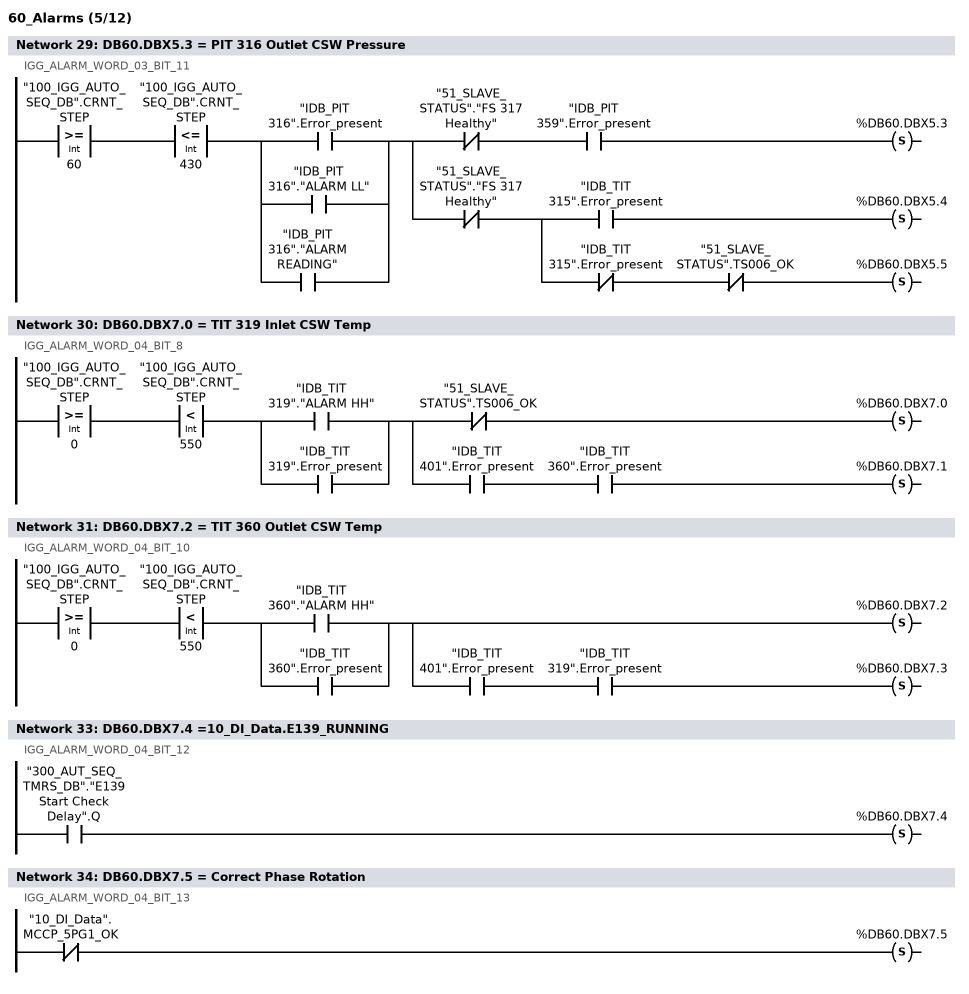
   RUNG wire#powerrail
      { S7_Templates := "SrcType := Int" } GE_Contact(in1 := "100_IGG_AUTO_SEQ_DB".CRNT_STEP, in2 := 60)
      { S7_Templates := "SrcType := Int" } LE_Contact(in1 := "100_IGG_AUTO_SEQ_DB".CRNT_STEP, in2 := 430)
      wire#w1
      Contact( "IDB_PIT 316".Error_present )
      wire#w2
      I_Contact( "51_SLAVE_STATUS"."FS 317 Healthy" )
      Contact( "IDB_PIT 359".Error_present )
      S_Coil( %DB60.DBX5.3 )
   END_RUNG
   RUNG wire#w1
      Contact( "IDB_PIT 316"."ALARM LL" )
   END_RUNG wire#w2
   RUNG wire#w1
      Contact( "IDB_PIT 316"."ALARM READING" )
   END_RUNG wire#w2
   RUNG wire#w2
      I_Contact( "51_SLAVE_STATUS"."FS 317 Healthy" )
      wire#w3
      Contact( "IDB_TIT 315".Error_present )
      S_Coil( %DB60.DBX5.4 )
   END_RUNG
   RUNG wire#w3
      I_Contact( "IDB_TIT 315".Error_present )
      I_Contact( "51_SLAVE_STATUS".TS006_OK )
      S_Coil( %DB60.DBX5.5 )
   END_RUNG
   // the same network as SCL:
   #_w1 := ("100_IGG_AUTO_SEQ_DB".CRNT_STEP >= 60) AND ("100_IGG_AUTO_SEQ_DB".CRNT_STEP <= 430) AND ("IDB_PIT 316".Error_present OR "IDB_PIT 316"."ALARM LL" OR "IDB_PIT 316"."ALARM READING");
   IF #_w1 AND NOT "51_SLAVE_STATUS"."FS 317 Healthy" AND "IDB_PIT 359".Error_present THEN
       %DB60.DBX5.3 := TRUE;
   END_IF;
   #_w2 := #_w1 AND NOT "51_SLAVE_STATUS"."FS 317 Healthy";
   IF #_w2 AND "IDB_TIT 315".Error_present THEN %DB60.DBX5.4 := TRUE; END_IF;
   IF #_w2 AND NOT "IDB_TIT 315".Error_present AND NOT "51_SLAVE_STATUS".TS006_OK THEN
       %DB60.DBX5.5 := TRUE;
   END_IF;
END_REGION

REGION Network 30: DB60.DBX7.0 = TIT 319 Inlet CSW Temp
   // IGG_ALARM_WORD_04_BIT_8
   RUNG wire#powerrail
      { S7_Templates := "SrcType := Int" } GE_Contact(in1 := "100_IGG_AUTO_SEQ_DB".CRNT_STEP, in2 := 0)
      { S7_Templates := "SrcType := Int" } LT_Contact(in1 := "100_IGG_AUTO_SEQ_DB".CRNT_STEP, in2 := 550)
      wire#w1
      Contact( "IDB_TIT 319"."ALARM HH" )
      wire#w2
      I_Contact( "51_SLAVE_STATUS".TS006_OK )
      S_Coil( %DB60.DBX7.0 )
   END_RUNG
   RUNG wire#w1
      Contact( "IDB_TIT 319".Error_present )
   END_RUNG wire#w2
   RUNG wire#w2
      Contact( "IDB_TIT 401".Error_present )
      Contact( "IDB_TIT 360".Error_present )
      S_Coil( %DB60.DBX7.1 )
   END_RUNG
   // the same network as SCL:
   #_w1 := ("100_IGG_AUTO_SEQ_DB".CRNT_STEP >= 0) AND ("100_IGG_AUTO_SEQ_DB".CRNT_STEP < 550) AND ("IDB_TIT 319"."ALARM HH" OR "IDB_TIT 319".Error_present);
   IF #_w1 AND NOT "51_SLAVE_STATUS".TS006_OK THEN %DB60.DBX7.0 := TRUE; END_IF;
   IF #_w1 AND "IDB_TIT 401".Error_present AND "IDB_TIT 360".Error_present THEN %DB60.DBX7.1 := TRUE; END_IF;
END_REGION

REGION Network 31: DB60.DBX7.2 = TIT 360 Outlet CSW Temp
   // IGG_ALARM_WORD_04_BIT_10
   RUNG wire#powerrail
      { S7_Templates := "SrcType := Int" } GE_Contact(in1 := "100_IGG_AUTO_SEQ_DB".CRNT_STEP, in2 := 0)
      { S7_Templates := "SrcType := Int" } LT_Contact(in1 := "100_IGG_AUTO_SEQ_DB".CRNT_STEP, in2 := 550)
      wire#w1
      Contact( "IDB_TIT 360"."ALARM HH" )
      wire#w2
      S_Coil( %DB60.DBX7.2 )
   END_RUNG
   RUNG wire#w1
      Contact( "IDB_TIT 360".Error_present )
   END_RUNG wire#w2
   RUNG wire#w2
      Contact( "IDB_TIT 401".Error_present )
      Contact( "IDB_TIT 319".Error_present )
      S_Coil( %DB60.DBX7.3 )
   END_RUNG
   // the same network as SCL:
   #_w1 := ("100_IGG_AUTO_SEQ_DB".CRNT_STEP >= 0) AND ("100_IGG_AUTO_SEQ_DB".CRNT_STEP < 550) AND ("IDB_TIT 360"."ALARM HH" OR "IDB_TIT 360".Error_present);
   IF #_w1 THEN %DB60.DBX7.2 := TRUE; END_IF;
   IF #_w1 AND "IDB_TIT 401".Error_present AND "IDB_TIT 319".Error_present THEN %DB60.DBX7.3 := TRUE; END_IF;
END_REGION

REGION Network 33: DB60.DBX7.4 =10_DI_Data.E139_RUNNING
   // IGG_ALARM_WORD_04_BIT_12
   RUNG wire#powerrail
      Contact( "300_AUT_SEQ_TMRS_DB"."E139 Start Check Delay".Q )
      S_Coil( %DB60.DBX7.4 )
   END_RUNG
   // the same network as SCL:
   IF "300_AUT_SEQ_TMRS_DB"."E139 Start Check Delay".Q THEN %DB60.DBX7.4 := TRUE; END_IF;
END_REGION

REGION Network 34: DB60.DBX7.5 = Correct Phase Rotation
   // IGG_ALARM_WORD_04_BIT_13
   RUNG wire#powerrail
      I_Contact( "10_DI_Data".MCCP_5PG1_OK )
      S_Coil( %DB60.DBX7.5 )
   END_RUNG
   // the same network as SCL:
   IF NOT "10_DI_Data".MCCP_5PG1_OK THEN %DB60.DBX7.5 := TRUE; END_IF;
END_REGION

REGION Network 36: DB60.DBX6.0 = CV311 Fault
   // IGG_ALARM_WORD_04_BIT_0
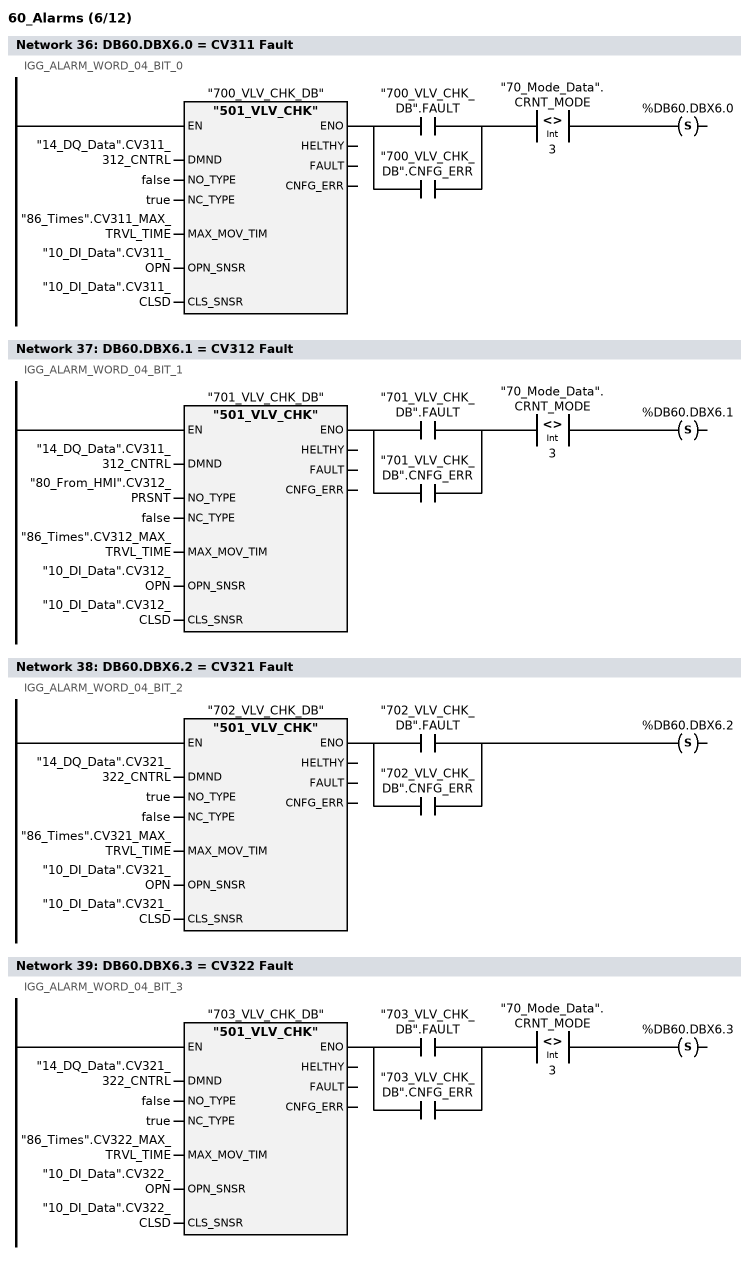
   RUNG wire#powerrail
      "700_VLV_CHK_DB"(DMND := "14_DQ_Data".CV311_312_CNTRL, NO_TYPE := false, NC_TYPE := true, MAX_MOV_TIM := "86_Times".CV311_MAX_TRVL_TIME, OPN_SNSR := "10_DI_Data".CV311_OPN, CLS_SNSR := "10_DI_Data".CV311_CLSD, HELTHY =>, FAULT =>, CNFG_ERR =>)
      wire#w1
      Contact( "700_VLV_CHK_DB".FAULT )
      wire#w2
      { S7_Templates := "SrcType := Int" } NE_Contact(in1 := "70_Mode_Data".CRNT_MODE, in2 := 3)
      S_Coil( %DB60.DBX6.0 )
   END_RUNG
   RUNG wire#w1
      Contact( "700_VLV_CHK_DB".CNFG_ERR )
   END_RUNG wire#w2
   // the same network as SCL:
   "700_VLV_CHK_DB"(DMND := "14_DQ_Data".CV311_312_CNTRL,   // "501_VLV_CHK"
                    NO_TYPE := false,
                    NC_TYPE := true,
                    MAX_MOV_TIM := "86_Times".CV311_MAX_TRVL_TIME,
                    OPN_SNSR := "10_DI_Data".CV311_OPN,
                    CLS_SNSR := "10_DI_Data".CV311_CLSD,
                    ENO => #_w1);
   IF #_w1 AND ("700_VLV_CHK_DB".FAULT OR "700_VLV_CHK_DB".CNFG_ERR) AND ("70_Mode_Data".CRNT_MODE <> 3) THEN
       %DB60.DBX6.0 := TRUE;
   END_IF;
END_REGION

REGION Network 37: DB60.DBX6.1 = CV312 Fault
   // IGG_ALARM_WORD_04_BIT_1
   RUNG wire#powerrail
      "701_VLV_CHK_DB"(DMND := "14_DQ_Data".CV311_312_CNTRL, NO_TYPE := "80_From_HMI".CV312_PRSNT, NC_TYPE := false, MAX_MOV_TIM := "86_Times".CV312_MAX_TRVL_TIME, OPN_SNSR := "10_DI_Data".CV312_OPN, CLS_SNSR := "10_DI_Data".CV312_CLSD, HELTHY =>, FAULT =>, CNFG_ERR =>)
      wire#w1
      Contact( "701_VLV_CHK_DB".FAULT )
      wire#w2
      { S7_Templates := "SrcType := Int" } NE_Contact(in1 := "70_Mode_Data".CRNT_MODE, in2 := 3)
      S_Coil( %DB60.DBX6.1 )
   END_RUNG
   RUNG wire#w1
      Contact( "701_VLV_CHK_DB".CNFG_ERR )
   END_RUNG wire#w2
   // the same network as SCL:
   "701_VLV_CHK_DB"(DMND := "14_DQ_Data".CV311_312_CNTRL,   // "501_VLV_CHK"
                    NO_TYPE := "80_From_HMI".CV312_PRSNT,
                    NC_TYPE := false,
                    MAX_MOV_TIM := "86_Times".CV312_MAX_TRVL_TIME,
                    OPN_SNSR := "10_DI_Data".CV312_OPN,
                    CLS_SNSR := "10_DI_Data".CV312_CLSD,
                    ENO => #_w1);
   IF #_w1 AND ("701_VLV_CHK_DB".FAULT OR "701_VLV_CHK_DB".CNFG_ERR) AND ("70_Mode_Data".CRNT_MODE <> 3) THEN
       %DB60.DBX6.1 := TRUE;
   END_IF;
END_REGION

REGION Network 38: DB60.DBX6.2 = CV321 Fault
   // IGG_ALARM_WORD_04_BIT_2
   RUNG wire#powerrail
      "702_VLV_CHK_DB"(DMND := "14_DQ_Data".CV321_322_CNTRL, NO_TYPE := true, NC_TYPE := false, MAX_MOV_TIM := "86_Times".CV321_MAX_TRVL_TIME, OPN_SNSR := "10_DI_Data".CV321_OPN, CLS_SNSR := "10_DI_Data".CV321_CLSD, HELTHY =>, FAULT =>, CNFG_ERR =>)
      wire#w1
      Contact( "702_VLV_CHK_DB".FAULT )
      wire#w2
      S_Coil( %DB60.DBX6.2 )
   END_RUNG
   RUNG wire#w1
      Contact( "702_VLV_CHK_DB".CNFG_ERR )
   END_RUNG wire#w2
   // the same network as SCL:
   "702_VLV_CHK_DB"(DMND := "14_DQ_Data".CV321_322_CNTRL,   // "501_VLV_CHK"
                    NO_TYPE := true,
                    NC_TYPE := false,
                    MAX_MOV_TIM := "86_Times".CV321_MAX_TRVL_TIME,
                    OPN_SNSR := "10_DI_Data".CV321_OPN,
                    CLS_SNSR := "10_DI_Data".CV321_CLSD,
                    ENO => #_w1);
   IF #_w1 AND ("702_VLV_CHK_DB".FAULT OR "702_VLV_CHK_DB".CNFG_ERR) THEN %DB60.DBX6.2 := TRUE; END_IF;
END_REGION

REGION Network 39: DB60.DBX6.3 = CV322 Fault
   // IGG_ALARM_WORD_04_BIT_3
   RUNG wire#powerrail
      "703_VLV_CHK_DB"(DMND := "14_DQ_Data".CV321_322_CNTRL, NO_TYPE := false, NC_TYPE := true, MAX_MOV_TIM := "86_Times".CV322_MAX_TRVL_TIME, OPN_SNSR := "10_DI_Data".CV322_OPN, CLS_SNSR := "10_DI_Data".CV322_CLSD, HELTHY =>, FAULT =>, CNFG_ERR =>)
      wire#w1
      Contact( "703_VLV_CHK_DB".FAULT )
      wire#w2
      { S7_Templates := "SrcType := Int" } NE_Contact(in1 := "70_Mode_Data".CRNT_MODE, in2 := 3)
      S_Coil( %DB60.DBX6.3 )
   END_RUNG
   RUNG wire#w1
      Contact( "703_VLV_CHK_DB".CNFG_ERR )
   END_RUNG wire#w2
   // the same network as SCL:
   "703_VLV_CHK_DB"(DMND := "14_DQ_Data".CV321_322_CNTRL,   // "501_VLV_CHK"
                    NO_TYPE := false,
                    NC_TYPE := true,
                    MAX_MOV_TIM := "86_Times".CV322_MAX_TRVL_TIME,
                    OPN_SNSR := "10_DI_Data".CV322_OPN,
                    CLS_SNSR := "10_DI_Data".CV322_CLSD,
                    ENO => #_w1);
   IF #_w1 AND ("703_VLV_CHK_DB".FAULT OR "703_VLV_CHK_DB".CNFG_ERR) AND ("70_Mode_Data".CRNT_MODE <> 3) THEN
       %DB60.DBX6.3 := TRUE;
   END_IF;
END_REGION

REGION Network 40: DB60.DBX6.4 = CV401 Fault
   // IGG_ALARM_WORD_04_BIT_4
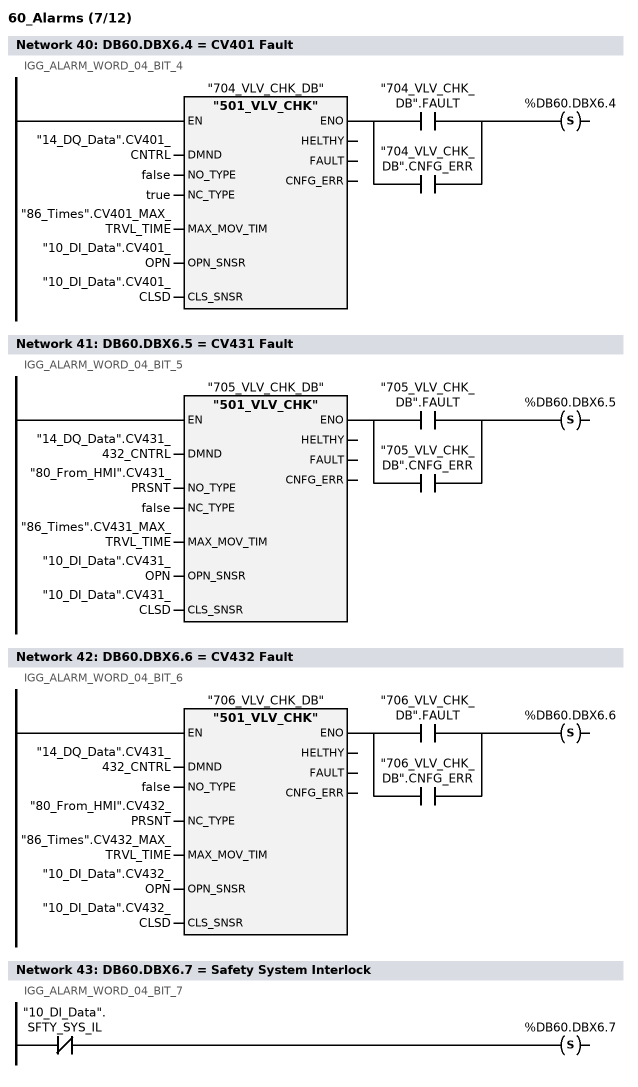
   RUNG wire#powerrail
      "704_VLV_CHK_DB"(DMND := "14_DQ_Data".CV401_CNTRL, NO_TYPE := false, NC_TYPE := true, MAX_MOV_TIM := "86_Times".CV401_MAX_TRVL_TIME, OPN_SNSR := "10_DI_Data".CV401_OPN, CLS_SNSR := "10_DI_Data".CV401_CLSD, HELTHY =>, FAULT =>, CNFG_ERR =>)
      wire#w1
      Contact( "704_VLV_CHK_DB".FAULT )
      wire#w2
      S_Coil( %DB60.DBX6.4 )
   END_RUNG
   RUNG wire#w1
      Contact( "704_VLV_CHK_DB".CNFG_ERR )
   END_RUNG wire#w2
   // the same network as SCL:
   "704_VLV_CHK_DB"(DMND := "14_DQ_Data".CV401_CNTRL,   // "501_VLV_CHK"
                    NO_TYPE := false,
                    NC_TYPE := true,
                    MAX_MOV_TIM := "86_Times".CV401_MAX_TRVL_TIME,
                    OPN_SNSR := "10_DI_Data".CV401_OPN,
                    CLS_SNSR := "10_DI_Data".CV401_CLSD,
                    ENO => #_w1);
   IF #_w1 AND ("704_VLV_CHK_DB".FAULT OR "704_VLV_CHK_DB".CNFG_ERR) THEN %DB60.DBX6.4 := TRUE; END_IF;
END_REGION

REGION Network 41: DB60.DBX6.5 = CV431 Fault
   // IGG_ALARM_WORD_04_BIT_5
   RUNG wire#powerrail
      "705_VLV_CHK_DB"(DMND := "14_DQ_Data".CV431_432_CNTRL, NO_TYPE := "80_From_HMI".CV431_PRSNT, NC_TYPE := false, MAX_MOV_TIM := "86_Times".CV431_MAX_TRVL_TIME, OPN_SNSR := "10_DI_Data".CV431_OPN, CLS_SNSR := "10_DI_Data".CV431_CLSD, HELTHY =>, FAULT =>, CNFG_ERR =>)
      wire#w1
      Contact( "705_VLV_CHK_DB".FAULT )
      wire#w2
      S_Coil( %DB60.DBX6.5 )
   END_RUNG
   RUNG wire#w1
      Contact( "705_VLV_CHK_DB".CNFG_ERR )
   END_RUNG wire#w2
   // the same network as SCL:
   "705_VLV_CHK_DB"(DMND := "14_DQ_Data".CV431_432_CNTRL,   // "501_VLV_CHK"
                    NO_TYPE := "80_From_HMI".CV431_PRSNT,
                    NC_TYPE := false,
                    MAX_MOV_TIM := "86_Times".CV431_MAX_TRVL_TIME,
                    OPN_SNSR := "10_DI_Data".CV431_OPN,
                    CLS_SNSR := "10_DI_Data".CV431_CLSD,
                    ENO => #_w1);
   IF #_w1 AND ("705_VLV_CHK_DB".FAULT OR "705_VLV_CHK_DB".CNFG_ERR) THEN %DB60.DBX6.5 := TRUE; END_IF;
END_REGION

REGION Network 42: DB60.DBX6.6 = CV432 Fault
   // IGG_ALARM_WORD_04_BIT_6
   RUNG wire#powerrail
      "706_VLV_CHK_DB"(DMND := "14_DQ_Data".CV431_432_CNTRL, NO_TYPE := false, NC_TYPE := "80_From_HMI".CV432_PRSNT, MAX_MOV_TIM := "86_Times".CV432_MAX_TRVL_TIME, OPN_SNSR := "10_DI_Data".CV432_OPN, CLS_SNSR := "10_DI_Data".CV432_CLSD, HELTHY =>, FAULT =>, CNFG_ERR =>)
      wire#w1
      Contact( "706_VLV_CHK_DB".FAULT )
      wire#w2
      S_Coil( %DB60.DBX6.6 )
   END_RUNG
   RUNG wire#w1
      Contact( "706_VLV_CHK_DB".CNFG_ERR )
   END_RUNG wire#w2
   // the same network as SCL:
   "706_VLV_CHK_DB"(DMND := "14_DQ_Data".CV431_432_CNTRL,   // "501_VLV_CHK"
                    NO_TYPE := false,
                    NC_TYPE := "80_From_HMI".CV432_PRSNT,
                    MAX_MOV_TIM := "86_Times".CV432_MAX_TRVL_TIME,
                    OPN_SNSR := "10_DI_Data".CV432_OPN,
                    CLS_SNSR := "10_DI_Data".CV432_CLSD,
                    ENO => #_w1);
   IF #_w1 AND ("706_VLV_CHK_DB".FAULT OR "706_VLV_CHK_DB".CNFG_ERR) THEN %DB60.DBX6.6 := TRUE; END_IF;
END_REGION

REGION Network 43: DB60.DBX6.7 = Safety System Interlock
   // IGG_ALARM_WORD_04_BIT_7
   RUNG wire#powerrail
      I_Contact( "10_DI_Data".SFTY_SYS_IL )
      S_Coil( %DB60.DBX6.7 )
   END_RUNG
   // the same network as SCL:
   IF NOT "10_DI_Data".SFTY_SYS_IL THEN %DB60.DBX6.7 := TRUE; END_IF;
END_REGION

REGION Network 45: New Alarm Check
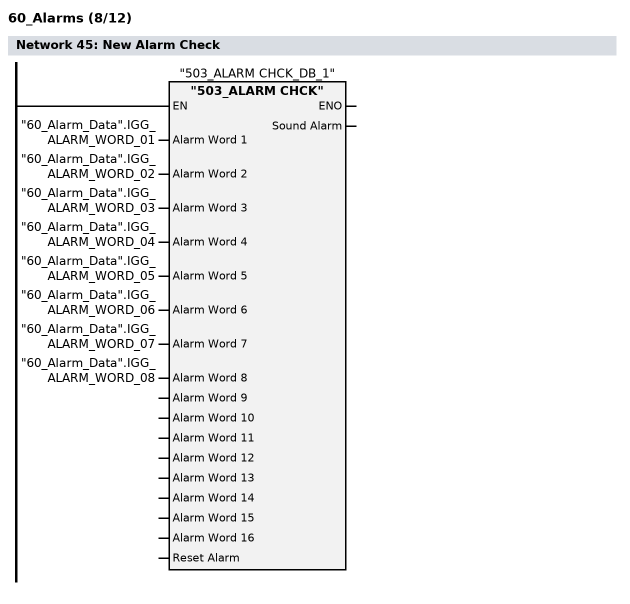
   RUNG wire#powerrail
      "503_ALARM CHCK_DB_1"("Alarm Word 1" := "60_Alarm_Data".IGG_ALARM_WORD_01, "Alarm Word 2" := "60_Alarm_Data".IGG_ALARM_WORD_02, "Alarm Word 3" := "60_Alarm_Data".IGG_ALARM_WORD_03, "Alarm Word 4" := "60_Alarm_Data".IGG_ALARM_WORD_04, "Alarm Word 5" := "60_Alarm_Data".IGG_ALARM_WORD_05, "Alarm Word 6" := "60_Alarm_Data".IGG_ALARM_WORD_06, "Alarm Word 7" := "60_Alarm_Data".IGG_ALARM_WORD_07, "Alarm Word 8" := "60_Alarm_Data".IGG_ALARM_WORD_08, "Alarm Word 9" :=, "Alarm Word 10" :=, "Alarm Word 11" :=, "Alarm Word 12" :=, "Alarm Word 13" :=, "Alarm Word 14" :=, "Alarm Word 15" :=, "Alarm Word 16" :=, "Reset Alarm" :=, "Sound Alarm" =>)
   END_RUNG
   // the same network as SCL:
   "503_ALARM CHCK_DB_1"("Alarm Word 1" := "60_Alarm_Data".IGG_ALARM_WORD_01,   // "503_ALARM CHCK"
                         "Alarm Word 2" := "60_Alarm_Data".IGG_ALARM_WORD_02,
                         "Alarm Word 3" := "60_Alarm_Data".IGG_ALARM_WORD_03,
                         "Alarm Word 4" := "60_Alarm_Data".IGG_ALARM_WORD_04,
                         "Alarm Word 5" := "60_Alarm_Data".IGG_ALARM_WORD_05,
                         "Alarm Word 6" := "60_Alarm_Data".IGG_ALARM_WORD_06,
                         "Alarm Word 7" := "60_Alarm_Data".IGG_ALARM_WORD_07,
                         "Alarm Word 8" := "60_Alarm_Data".IGG_ALARM_WORD_08);
END_REGION

REGION Network 46: Alarm reset
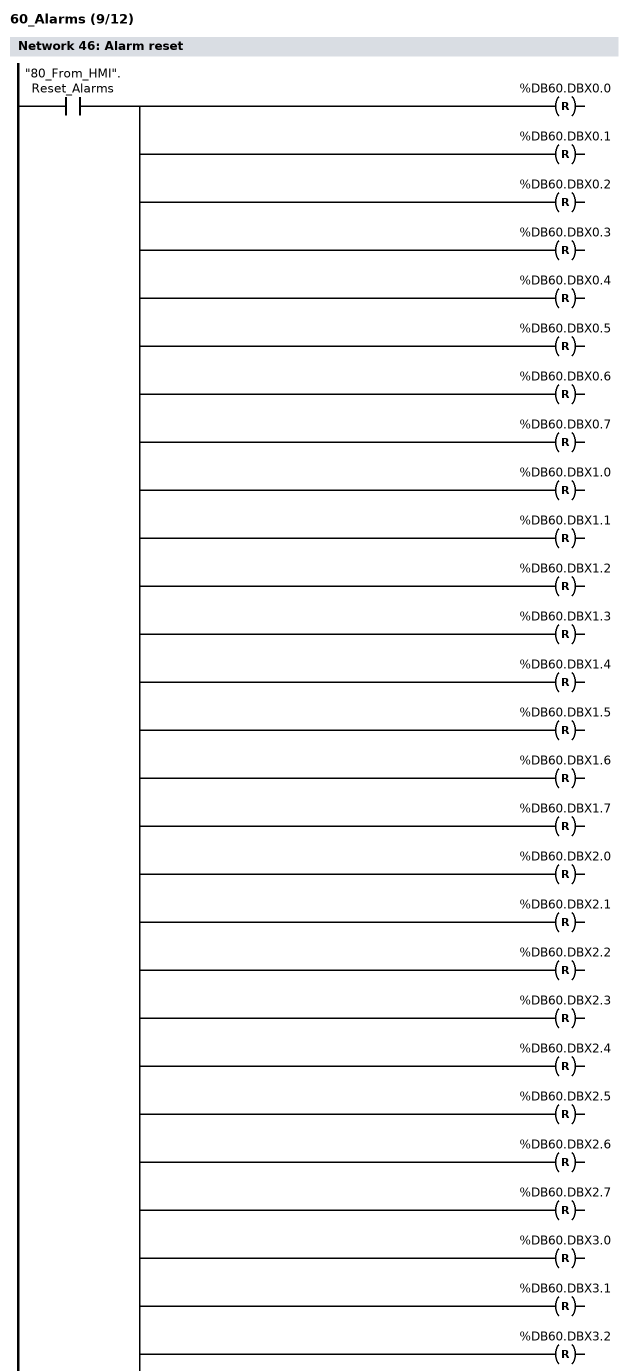
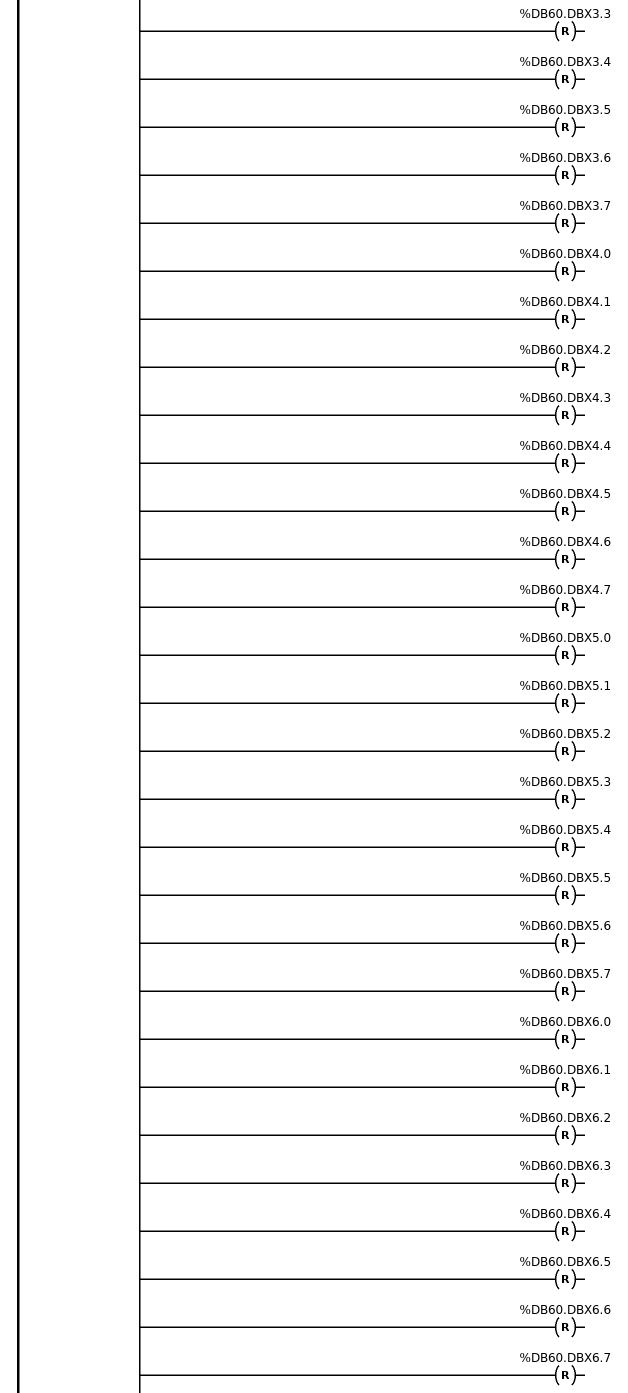
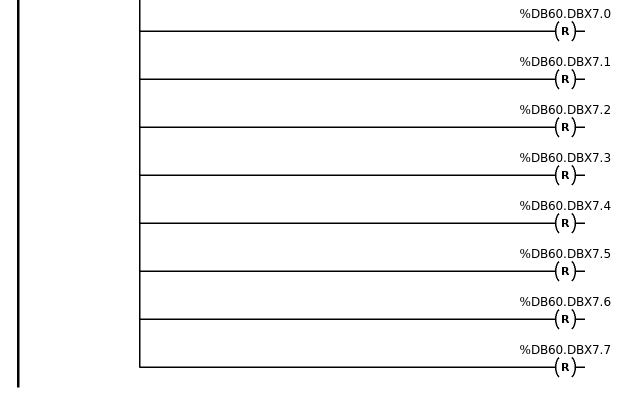
   RUNG wire#powerrail
      Contact( "80_From_HMI".Reset_Alarms )
      wire#w1
      R_Coil( %DB60.DBX0.0 )
   END_RUNG
   RUNG wire#w1
      R_Coil( %DB60.DBX0.1 )
   END_RUNG
   RUNG wire#w1
      R_Coil( %DB60.DBX0.2 )
   END_RUNG
   RUNG wire#w1
      R_Coil( %DB60.DBX0.3 )
   END_RUNG
   RUNG wire#w1
      R_Coil( %DB60.DBX0.4 )
   END_RUNG
   RUNG wire#w1
      R_Coil( %DB60.DBX0.5 )
   END_RUNG
   RUNG wire#w1
      R_Coil( %DB60.DBX0.6 )
   END_RUNG
   RUNG wire#w1
      R_Coil( %DB60.DBX0.7 )
   END_RUNG
   RUNG wire#w1
      R_Coil( %DB60.DBX1.0 )
   END_RUNG
   RUNG wire#w1
      R_Coil( %DB60.DBX1.1 )
   END_RUNG
   RUNG wire#w1
      R_Coil( %DB60.DBX1.2 )
   END_RUNG
   RUNG wire#w1
      R_Coil( %DB60.DBX1.3 )
   END_RUNG
   RUNG wire#w1
      R_Coil( %DB60.DBX1.4 )
   END_RUNG
   RUNG wire#w1
      R_Coil( %DB60.DBX1.5 )
   END_RUNG
   RUNG wire#w1
      R_Coil( %DB60.DBX1.6 )
   END_RUNG
   RUNG wire#w1
      R_Coil( %DB60.DBX1.7 )
   END_RUNG
   RUNG wire#w1
      R_Coil( %DB60.DBX2.0 )
   END_RUNG
   RUNG wire#w1
      R_Coil( %DB60.DBX2.1 )
   END_RUNG
   RUNG wire#w1
      R_Coil( %DB60.DBX2.2 )
   END_RUNG
   RUNG wire#w1
      R_Coil( %DB60.DBX2.3 )
   END_RUNG
   RUNG wire#w1
      R_Coil( %DB60.DBX2.4 )
   END_RUNG
   RUNG wire#w1
      R_Coil( %DB60.DBX2.5 )
   END_RUNG
   RUNG wire#w1
      R_Coil( %DB60.DBX2.6 )
   END_RUNG
   RUNG wire#w1
      R_Coil( %DB60.DBX2.7 )
   END_RUNG
   RUNG wire#w1
      R_Coil( %DB60.DBX3.0 )
   END_RUNG
   RUNG wire#w1
      R_Coil( %DB60.DBX3.1 )
   END_RUNG
   RUNG wire#w1
      R_Coil( %DB60.DBX3.2 )
   END_RUNG
   RUNG wire#w1
      R_Coil( %DB60.DBX3.3 )
   END_RUNG
   RUNG wire#w1
      R_Coil( %DB60.DBX3.4 )
   END_RUNG
   RUNG wire#w1
      R_Coil( %DB60.DBX3.5 )
   END_RUNG
   RUNG wire#w1
      R_Coil( %DB60.DBX3.6 )
   END_RUNG
   RUNG wire#w1
      R_Coil( %DB60.DBX3.7 )
   END_RUNG
   RUNG wire#w1
      R_Coil( %DB60.DBX4.0 )
   END_RUNG
   RUNG wire#w1
      R_Coil( %DB60.DBX4.1 )
   END_RUNG
   RUNG wire#w1
      R_Coil( %DB60.DBX4.2 )
   END_RUNG
   RUNG wire#w1
      R_Coil( %DB60.DBX4.3 )
   END_RUNG
   RUNG wire#w1
      R_Coil( %DB60.DBX4.4 )
   END_RUNG
   RUNG wire#w1
      R_Coil( %DB60.DBX4.5 )
   END_RUNG
   RUNG wire#w1
      R_Coil( %DB60.DBX4.6 )
   END_RUNG
   RUNG wire#w1
      R_Coil( %DB60.DBX4.7 )
   END_RUNG
   RUNG wire#w1
      R_Coil( %DB60.DBX5.0 )
   END_RUNG
   RUNG wire#w1
      R_Coil( %DB60.DBX5.1 )
   END_RUNG
   RUNG wire#w1
      R_Coil( %DB60.DBX5.2 )
   END_RUNG
   RUNG wire#w1
      R_Coil( %DB60.DBX5.3 )
   END_RUNG
   RUNG wire#w1
      R_Coil( %DB60.DBX5.4 )
   END_RUNG
   RUNG wire#w1
      R_Coil( %DB60.DBX5.5 )
   END_RUNG
   RUNG wire#w1
      R_Coil( %DB60.DBX5.6 )
   END_RUNG
   RUNG wire#w1
      R_Coil( %DB60.DBX5.7 )
   END_RUNG
   RUNG wire#w1
      R_Coil( %DB60.DBX6.0 )
   END_RUNG
   RUNG wire#w1
      R_Coil( %DB60.DBX6.1 )
   END_RUNG
   RUNG wire#w1
      R_Coil( %DB60.DBX6.2 )
   END_RUNG
   RUNG wire#w1
      R_Coil( %DB60.DBX6.3 )
   END_RUNG
   RUNG wire#w1
      R_Coil( %DB60.DBX6.4 )
   END_RUNG
   RUNG wire#w1
      R_Coil( %DB60.DBX6.5 )
   END_RUNG
   RUNG wire#w1
      R_Coil( %DB60.DBX6.6 )
   END_RUNG
   RUNG wire#w1
      R_Coil( %DB60.DBX6.7 )
   END_RUNG
   RUNG wire#w1
      R_Coil( %DB60.DBX7.0 )
   END_RUNG
   RUNG wire#w1
      R_Coil( %DB60.DBX7.1 )
   END_RUNG
   RUNG wire#w1
      R_Coil( %DB60.DBX7.2 )
   END_RUNG
   RUNG wire#w1
      R_Coil( %DB60.DBX7.3 )
   END_RUNG
   RUNG wire#w1
      R_Coil( %DB60.DBX7.4 )
   END_RUNG
   RUNG wire#w1
      R_Coil( %DB60.DBX7.5 )
   END_RUNG
   RUNG wire#w1
      R_Coil( %DB60.DBX7.6 )
   END_RUNG
   RUNG wire#w1
      R_Coil( %DB60.DBX7.7 )
   END_RUNG
   // the same network as SCL:
   IF "80_From_HMI".Reset_Alarms THEN
       %DB60.DBX0.0 := FALSE;
       %DB60.DBX0.1 := FALSE;
       %DB60.DBX0.2 := FALSE;
       %DB60.DBX0.3 := FALSE;
       %DB60.DBX0.4 := FALSE;
       %DB60.DBX0.5 := FALSE;
       %DB60.DBX0.6 := FALSE;
       %DB60.DBX0.7 := FALSE;
       %DB60.DBX1.0 := FALSE;
       %DB60.DBX1.1 := FALSE;
       %DB60.DBX1.2 := FALSE;
       %DB60.DBX1.3 := FALSE;
       %DB60.DBX1.4 := FALSE;
       %DB60.DBX1.5 := FALSE;
       %DB60.DBX1.6 := FALSE;
       %DB60.DBX1.7 := FALSE;
       %DB60.DBX2.0 := FALSE;
       %DB60.DBX2.1 := FALSE;
       %DB60.DBX2.2 := FALSE;
       %DB60.DBX2.3 := FALSE;
       %DB60.DBX2.4 := FALSE;
       %DB60.DBX2.5 := FALSE;
       %DB60.DBX2.6 := FALSE;
       %DB60.DBX2.7 := FALSE;
       %DB60.DBX3.0 := FALSE;
       %DB60.DBX3.1 := FALSE;
       %DB60.DBX3.2 := FALSE;
       %DB60.DBX3.3 := FALSE;
       %DB60.DBX3.4 := FALSE;
       %DB60.DBX3.5 := FALSE;
       %DB60.DBX3.6 := FALSE;
       %DB60.DBX3.7 := FALSE;
       %DB60.DBX4.0 := FALSE;
       %DB60.DBX4.1 := FALSE;
       %DB60.DBX4.2 := FALSE;
       %DB60.DBX4.3 := FALSE;
       %DB60.DBX4.4 := FALSE;
       %DB60.DBX4.5 := FALSE;
       %DB60.DBX4.6 := FALSE;
       %DB60.DBX4.7 := FALSE;
       %DB60.DBX5.0 := FALSE;
       %DB60.DBX5.1 := FALSE;
       %DB60.DBX5.2 := FALSE;
       %DB60.DBX5.3 := FALSE;
       %DB60.DBX5.4 := FALSE;
       %DB60.DBX5.5 := FALSE;
       %DB60.DBX5.6 := FALSE;
       %DB60.DBX5.7 := FALSE;
       %DB60.DBX6.0 := FALSE;
       %DB60.DBX6.1 := FALSE;
       %DB60.DBX6.2 := FALSE;
       %DB60.DBX6.3 := FALSE;
       %DB60.DBX6.4 := FALSE;
       %DB60.DBX6.5 := FALSE;
       %DB60.DBX6.6 := FALSE;
       %DB60.DBX6.7 := FALSE;
       %DB60.DBX7.0 := FALSE;
       %DB60.DBX7.1 := FALSE;
       %DB60.DBX7.2 := FALSE;
       %DB60.DBX7.3 := FALSE;
       %DB60.DBX7.4 := FALSE;
       %DB60.DBX7.5 := FALSE;
       %DB60.DBX7.6 := FALSE;
       %DB60.DBX7.7 := FALSE;
   END_IF;
END_REGION

REGION Network 47: Alarm reset II
   // testing
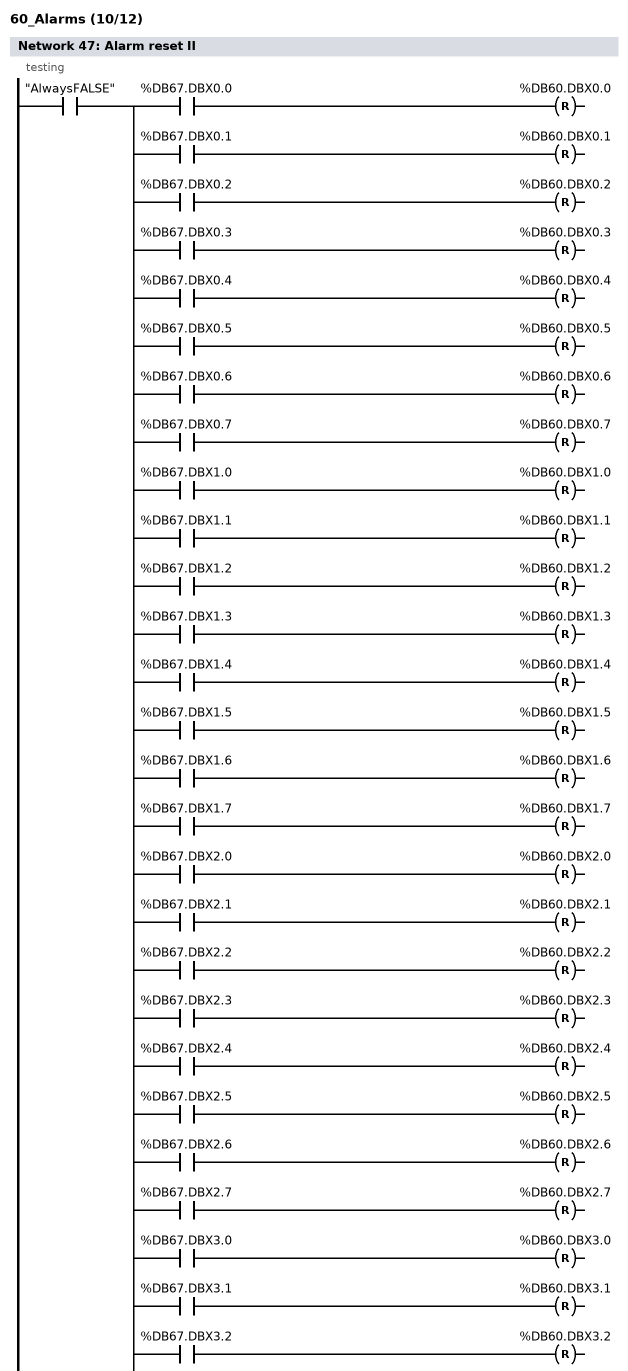
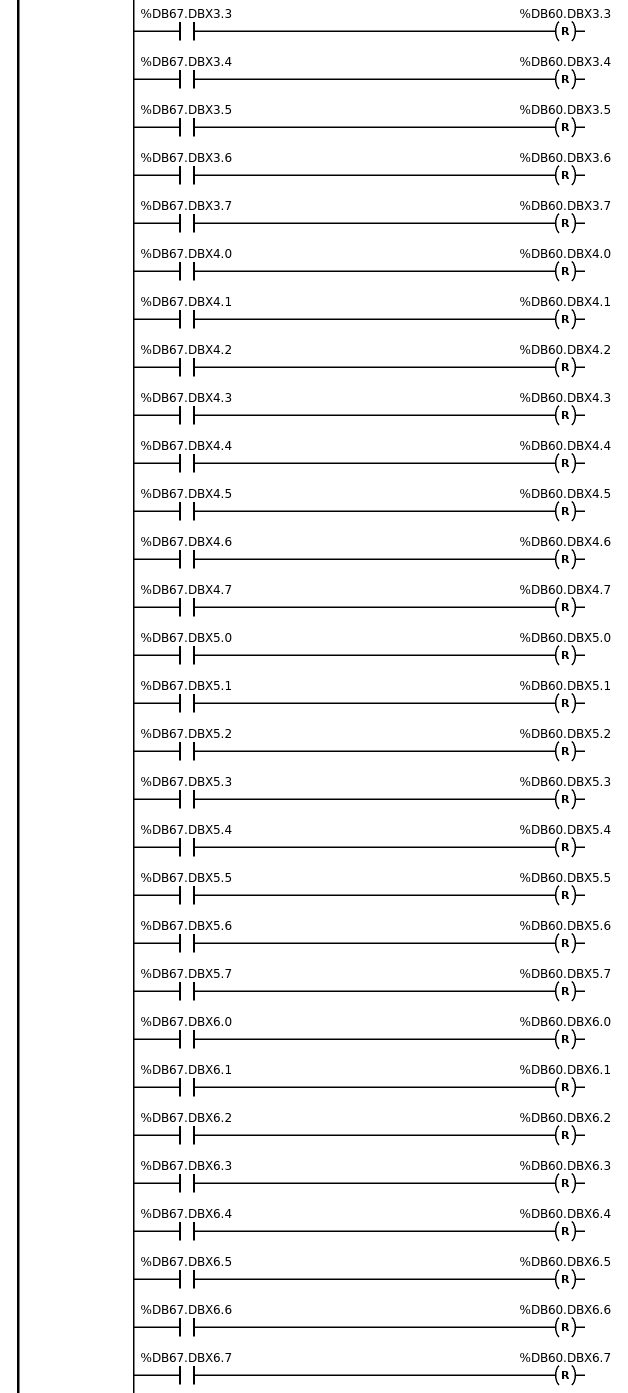
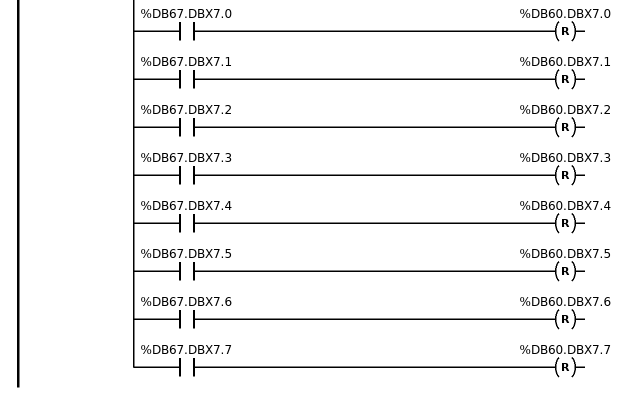
   RUNG wire#powerrail
      Contact( "AlwaysFALSE" )
      wire#w1
      Contact( %DB67.DBX0.0 )
      R_Coil( %DB60.DBX0.0 )
   END_RUNG
   RUNG wire#w1
      Contact( %DB67.DBX0.1 )
      R_Coil( %DB60.DBX0.1 )
   END_RUNG
   RUNG wire#w1
      Contact( %DB67.DBX0.2 )
      R_Coil( %DB60.DBX0.2 )
   END_RUNG
   RUNG wire#w1
      Contact( %DB67.DBX0.3 )
      R_Coil( %DB60.DBX0.3 )
   END_RUNG
   RUNG wire#w1
      Contact( %DB67.DBX0.4 )
      R_Coil( %DB60.DBX0.4 )
   END_RUNG
   RUNG wire#w1
      Contact( %DB67.DBX0.5 )
      R_Coil( %DB60.DBX0.5 )
   END_RUNG
   RUNG wire#w1
      Contact( %DB67.DBX0.6 )
      R_Coil( %DB60.DBX0.6 )
   END_RUNG
   RUNG wire#w1
      Contact( %DB67.DBX0.7 )
      R_Coil( %DB60.DBX0.7 )
   END_RUNG
   RUNG wire#w1
      Contact( %DB67.DBX1.0 )
      R_Coil( %DB60.DBX1.0 )
   END_RUNG
   RUNG wire#w1
      Contact( %DB67.DBX1.1 )
      R_Coil( %DB60.DBX1.1 )
   END_RUNG
   RUNG wire#w1
      Contact( %DB67.DBX1.2 )
      R_Coil( %DB60.DBX1.2 )
   END_RUNG
   RUNG wire#w1
      Contact( %DB67.DBX1.3 )
      R_Coil( %DB60.DBX1.3 )
   END_RUNG
   RUNG wire#w1
      Contact( %DB67.DBX1.4 )
      R_Coil( %DB60.DBX1.4 )
   END_RUNG
   RUNG wire#w1
      Contact( %DB67.DBX1.5 )
      R_Coil( %DB60.DBX1.5 )
   END_RUNG
   RUNG wire#w1
      Contact( %DB67.DBX1.6 )
      R_Coil( %DB60.DBX1.6 )
   END_RUNG
   RUNG wire#w1
      Contact( %DB67.DBX1.7 )
      R_Coil( %DB60.DBX1.7 )
   END_RUNG
   RUNG wire#w1
      Contact( %DB67.DBX2.0 )
      R_Coil( %DB60.DBX2.0 )
   END_RUNG
   RUNG wire#w1
      Contact( %DB67.DBX2.1 )
      R_Coil( %DB60.DBX2.1 )
   END_RUNG
   RUNG wire#w1
      Contact( %DB67.DBX2.2 )
      R_Coil( %DB60.DBX2.2 )
   END_RUNG
   RUNG wire#w1
      Contact( %DB67.DBX2.3 )
      R_Coil( %DB60.DBX2.3 )
   END_RUNG
   RUNG wire#w1
      Contact( %DB67.DBX2.4 )
      R_Coil( %DB60.DBX2.4 )
   END_RUNG
   RUNG wire#w1
      Contact( %DB67.DBX2.5 )
      R_Coil( %DB60.DBX2.5 )
   END_RUNG
   RUNG wire#w1
      Contact( %DB67.DBX2.6 )
      R_Coil( %DB60.DBX2.6 )
   END_RUNG
   RUNG wire#w1
      Contact( %DB67.DBX2.7 )
      R_Coil( %DB60.DBX2.7 )
   END_RUNG
   RUNG wire#w1
      Contact( %DB67.DBX3.0 )
      R_Coil( %DB60.DBX3.0 )
   END_RUNG
   RUNG wire#w1
      Contact( %DB67.DBX3.1 )
      R_Coil( %DB60.DBX3.1 )
   END_RUNG
   RUNG wire#w1
      Contact( %DB67.DBX3.2 )
      R_Coil( %DB60.DBX3.2 )
   END_RUNG
   RUNG wire#w1
      Contact( %DB67.DBX3.3 )
      R_Coil( %DB60.DBX3.3 )
   END_RUNG
   RUNG wire#w1
      Contact( %DB67.DBX3.4 )
      R_Coil( %DB60.DBX3.4 )
   END_RUNG
   RUNG wire#w1
      Contact( %DB67.DBX3.5 )
      R_Coil( %DB60.DBX3.5 )
   END_RUNG
   RUNG wire#w1
      Contact( %DB67.DBX3.6 )
      R_Coil( %DB60.DBX3.6 )
   END_RUNG
   RUNG wire#w1
      Contact( %DB67.DBX3.7 )
      R_Coil( %DB60.DBX3.7 )
   END_RUNG
   RUNG wire#w1
      Contact( %DB67.DBX4.0 )
      R_Coil( %DB60.DBX4.0 )
   END_RUNG
   RUNG wire#w1
      Contact( %DB67.DBX4.1 )
      R_Coil( %DB60.DBX4.1 )
   END_RUNG
   RUNG wire#w1
      Contact( %DB67.DBX4.2 )
      R_Coil( %DB60.DBX4.2 )
   END_RUNG
   RUNG wire#w1
      Contact( %DB67.DBX4.3 )
      R_Coil( %DB60.DBX4.3 )
   END_RUNG
   RUNG wire#w1
      Contact( %DB67.DBX4.4 )
      R_Coil( %DB60.DBX4.4 )
   END_RUNG
   RUNG wire#w1
      Contact( %DB67.DBX4.5 )
      R_Coil( %DB60.DBX4.5 )
   END_RUNG
   RUNG wire#w1
      Contact( %DB67.DBX4.6 )
      R_Coil( %DB60.DBX4.6 )
   END_RUNG
   RUNG wire#w1
      Contact( %DB67.DBX4.7 )
      R_Coil( %DB60.DBX4.7 )
   END_RUNG
   RUNG wire#w1
      Contact( %DB67.DBX5.0 )
      R_Coil( %DB60.DBX5.0 )
   END_RUNG
   RUNG wire#w1
      Contact( %DB67.DBX5.1 )
      R_Coil( %DB60.DBX5.1 )
   END_RUNG
   RUNG wire#w1
      Contact( %DB67.DBX5.2 )
      R_Coil( %DB60.DBX5.2 )
   END_RUNG
   RUNG wire#w1
      Contact( %DB67.DBX5.3 )
      R_Coil( %DB60.DBX5.3 )
   END_RUNG
   RUNG wire#w1
      Contact( %DB67.DBX5.4 )
      R_Coil( %DB60.DBX5.4 )
   END_RUNG
   RUNG wire#w1
      Contact( %DB67.DBX5.5 )
      R_Coil( %DB60.DBX5.5 )
   END_RUNG
   RUNG wire#w1
      Contact( %DB67.DBX5.6 )
      R_Coil( %DB60.DBX5.6 )
   END_RUNG
   RUNG wire#w1
      Contact( %DB67.DBX5.7 )
      R_Coil( %DB60.DBX5.7 )
   END_RUNG
   RUNG wire#w1
      Contact( %DB67.DBX6.0 )
      R_Coil( %DB60.DBX6.0 )
   END_RUNG
   RUNG wire#w1
      Contact( %DB67.DBX6.1 )
      R_Coil( %DB60.DBX6.1 )
   END_RUNG
   RUNG wire#w1
      Contact( %DB67.DBX6.2 )
      R_Coil( %DB60.DBX6.2 )
   END_RUNG
   RUNG wire#w1
      Contact( %DB67.DBX6.3 )
      R_Coil( %DB60.DBX6.3 )
   END_RUNG
   RUNG wire#w1
      Contact( %DB67.DBX6.4 )
      R_Coil( %DB60.DBX6.4 )
   END_RUNG
   RUNG wire#w1
      Contact( %DB67.DBX6.5 )
      R_Coil( %DB60.DBX6.5 )
   END_RUNG
   RUNG wire#w1
      Contact( %DB67.DBX6.6 )
      R_Coil( %DB60.DBX6.6 )
   END_RUNG
   RUNG wire#w1
      Contact( %DB67.DBX6.7 )
      R_Coil( %DB60.DBX6.7 )
   END_RUNG
   RUNG wire#w1
      Contact( %DB67.DBX7.0 )
      R_Coil( %DB60.DBX7.0 )